
               REGION "FLASHING"
                   IF #retLogical.acutal.btn[#pBtn] THEN

                       REGION "FLASH COLOR 1"
                           IF NOT #btnParams.btn[#pBtn].flash THEN
                               IF #old.btnParam.btn[#pBtn].flash THEN
                                   #color := #btnParams.btn[#pBtn].cOn1;
                                   #draw := TRUE;
                               END_IF;
                           END_IF;
                       END_REGION

                       REGION "FLASH COLOR 2"
                           IF #btnParams.btn[#pBtn].flash THEN
                               IF NOT #old.btnParam.btn[#pBtn].flash THEN
                                   #color := #btnParams.btn[#pBtn].cOn2;
                                   #draw := TRUE;
                               END_IF;
                           END_IF;
                       END_REGION

                   END_IF;
               END_REGION

               REGION "DRAW TO BUTTON"
                   IF #draw THEN
                       #draw := FALSE;
                       "KP8 Driver: Color"(btnColor := #colorMask,
                                           btnNum := #pBtn,
                                           lblColor := #color);
                   END_IF;
               END_REGION

           END_FOR;
       END_REGION

   END_REGION

   REGION "CHANGE DETECTION"
       #old.btnParam := #btnParams;
       #old.kp8DI := #kp8DI;
       #old.logical := #retLogical.acutal;
       #old.physical := #btnPress;
   END_REGION

   REGION "OUTPUT"
       #kp8DQ := #colorMask;
       #physical := #retPhysical;
       #logical := #retLogical;
   END_REGION
END_FUNCTION_BLOCK

FUNCTION "KP8 Driver: HMI Emulator: Animation" : USInt   // FC26, SCL
{ S7_Optimized_Access := 'TRUE' }
VERSION : 0.1
   VAR_INPUT
      kp8Color : DWord;
      btnNumber : Int;
   END_VAR
   VAR_TEMP
      animate : USInt;
      blue : USInt;
      colorDWord : DWord;
      colorInt : DInt;
      green : USInt;
      off : USInt;
      red : USInt;
      white : USInt;
      yellow : USInt;
   END_VAR
   VAR CONSTANT
      blueMask : DInt := 16#0000_0100;
      btnMask : DInt := 16#0101_0100;
      greenMask : DInt := 16#0001_0000;
      offMask : DInt := 16#0000_0000;
      redMask : DInt := 16#0100_0000;
      whiteMask : DInt := 16#0101_0100;
      yellowMask : DInt := 16#0101_0000;
   END_VAR
BEGIN
   REGION "COPY TO LOCAL"
       #blue := "BLUE_LIGHT_BACKGROUND";
       #green := "GREEN_LIGHT_BACKGROUND";
       #off := "invisible";
       #red := "RED_LIGHT_BACKGROUND";
       #white := "WHITE_BACKGROUND";
       #yellow := "YELLOW_LIGHT_BACKGROUND";
   END_REGION

   REGION "ISOLATE BUTTON COLOR"
       #colorDWord := SHR_DWORD(IN := #kp8Color,N := INT_TO_ULINT(#btnNumber));
       #colorDWord := #colorDWord AND #btnMask;
       #colorInt := DWORD_TO_DINT(#colorDWord);
   END_REGION

   REGION "DETERMINE ANIMATION"
       CASE #colorInt OF
           #blueMask:
               #animate := #blue;
           #greenMask:
               #animate := #green;
           #redMask:
               #animate := #red;
           #whiteMask:
               #animate := #white;
           #yellowMask:
               #animate := #yellow;
           ELSE
               #animate := #off;
       END_CASE;
   END_REGION

   REGION "RETURN VALUE"
       #"KP8 Driver: HMI Emulator: Animation" := #animate;
   END_REGION
END_FUNCTION

FUNCTION "KP8 Driver: Group" : Void   // FC50, SCL
{ S7_Optimized_Access := 'TRUE' }
VERSION : 0.1
   VAR_INPUT
      btnNumber : Int;
      btnsParams : "KP8 Driver: Parameters: 8 Buttons";
   END_VAR
   VAR_IN_OUT
      logical : "KP8 Driver: Feedback Data";
   END_VAR
   VAR_TEMP
      pBtn : Int;
      retLogical : "KP8 Driver: Feedback Data";
      testGroup : Int;
      thisGroup : Int;
   END_VAR
BEGIN
   REGION "EXIT IF GROUP EQUALS 0"
       #thisGroup := #btnsParams.btn[#btnNumber].group;
       IF #thisGroup = 0 THEN
           RETURN;
       END_IF;
   END_REGION

   REGION "COPY TO LOCAL"
       #retLogical := #logical;
   END_REGION

   REGION "FOR EACH BUTTONS' PARAMETERS"
       FOR #pBtn := 0 TO 7 DO

           REGION "SKIP THE CURRENT BUTTON"
               IF #pBtn = #btnNumber THEN
                   GOTO NEXT;
               END_IF;
           END_REGION

           REGION "GROUP EXCLUSION"
               #testGroup := #btnsParams.btn[#pBtn].group;
               IF #testGroup = #thisGroup THEN
                   #retLogical.acutal.btn[#pBtn] := FALSE;
               END_IF;
           END_REGION

       NEXT:
           ;

       END_FOR;
   END_REGION

   REGION "OUTPUT"
       #logical := #retLogical;
   END_REGION
END_FUNCTION

FUNCTION "KP8 Driver: Toggle" : Void   // FC51, SCL
{ S7_Optimized_Access := 'TRUE' }
VERSION : 0.1
   VAR_INPUT
      signal : Bool;   // edge signal
   END_VAR
   VAR_IN_OUT
      state : Bool;   // logical button state
   END_VAR
BEGIN
   IF #signal THEN
       #state := NOT #state;
   END_IF;
END_FUNCTION

FUNCTION "KP8 Driver: Feedback" : Void   // FC52, SCL
{ S7_Optimized_Access := 'TRUE' }
VERSION : 0.1
   VAR_INPUT
      signal : Bool;
      oldSignal : Bool;
      btnNumber : Int;
   END_VAR
   VAR_IN_OUT
      feedback : "KP8 Driver: Feedback Data";
   END_VAR
   VAR_TEMP
      ret : "KP8 Driver: Feedback Data";
   END_VAR
BEGIN
   REGION "COPY TO LOCAL"
       #ret := #feedback;
       #ret.acutal.btn[#btnNumber] := #signal;
   END_REGION

   REGION "DEFAULT"
       #ret.rising.btn[#btnNumber] := FALSE;
       #ret.falling.btn[#btnNumber] := FALSE;
   END_REGION

   REGION "ON NEW INPUT"
       IF #signal <> #oldSignal THEN

           REGION "RISING EDGE"
               IF #signal AND NOT #oldSignal THEN
                   #ret.rising.btn[#btnNumber] := TRUE;
               END_IF;
           END_REGION

           REGION "FALLING EDGE"
               IF NOT #signal AND #oldSignal THEN
                   #ret.falling.btn[#btnNumber] := TRUE;
               END_IF;
           END_REGION

       END_IF;
   END_REGION


   REGION "OUTPUT"
       #feedback := #ret;
   END_REGION
END_FUNCTION

FUNCTION "KP8 Driver: State" : Void   // FC53, SCL
{ S7_Optimized_Access := 'TRUE' }
VERSION : 0.1
   VAR_INPUT
      press : "KP8 Driver: Feedback Data";
      btnNumber : Int;
      btnParams : "KP8 Driver: Parameters: 8 Buttons";
   END_VAR
   VAR_IN_OUT
      state : "KP8 Driver: Feedback Data";
   END_VAR
   VAR_TEMP
      pBtn : Int;
      retState : "KP8 Driver: Feedback Data";
   END_VAR
BEGIN
   REGION "RETURN ON INACTIVE BUTTON"
       IF NOT #btnParams.btn[#btnNumber].activate THEN
           RETURN;
       END_IF;
   END_REGION

   REGION "COPY TO LOCAL"
       #retState := #state;
   END_REGION

   REGION "MODE IS MOMENTARY"
       IF NOT #btnParams.btn[#btnNumber].mode THEN
           #retState.acutal.btn[#btnNumber] := #press.acutal.btn[#btnNumber];
       END_IF;
   END_REGION

   REGION "MAINTINED"
       IF #btnParams.btn[#btnNumber].mode THEN
           "KP8 Driver: Toggle"(signal := #press.rising.btn[#btnNumber],
                                state := #retState.acutal.btn[#btnNumber]);
       END_IF;
   END_REGION

   REGION "GROUP EXCLUSIVITY"
       IF #press.rising.btn[#btnNumber] THEN
           "KP8 Driver: Group"(btnNumber := #btnNumber,
                               btnsParams := #btnParams,
                               logical := #retState);
       END_IF;
   END_REGION

   REGION "OUTPUT"
       #state := #retState;
   END_REGION
END_FUNCTION

FUNCTION "KP8 Driver: Color" : Void   // FC54, SCL
{ S7_Optimized_Access := 'TRUE' }
VERSION : 0.1
   VAR_INPUT
      btnNum : Int;
      lblColor : String;   // 'red', 'green', 'blue', 'yellow', 'white', 'off'
   END_VAR
   VAR_IN_OUT
      btnColor : DWord;
   END_VAR
   VAR_TEMP
      btnMask : DWord;
      uColor : String;
      ret : DWord;
   END_VAR
   VAR CONSTANT
      btnMskRed : DWord := DWORD#16#0100_0000;
      btnMskGreen : DWord := DWORD#16#0001_0000;
      btnMskBlue : DWord := DWORD#16#0000_0100;
      btnMskYellow : DWord := DWORD#16#0101_0000;
      btnMskWhite : DWord := DWORD#16#0101_0100;
      btnMskOff : DWord := DWORD#16#FEFE_FEFF;
   END_VAR
BEGIN
   #ret := #btnColor;

   #ret := #ret AND ROL(IN := #btnMskOff,
                        N := INT_TO_UDINT(#btnNum));

   #uColor := #lblColor;
   "Upper"(#uColor);

   IF (#uColor = 'RED') THEN
       #btnMask := #btnMskRed;
   ELSIF (#uColor = 'GREEN') THEN
       #btnMask := #btnMskGreen;
   ELSIF (#uColor = 'BLUE') THEN
       #btnMask := #btnMskBlue;
   ELSIF (#uColor = 'YELLOW') THEN
       #btnMask := #btnMskYellow;
   ELSIF (#uColor = 'WHITE') THEN
       #btnMask := #btnMskWhite;
   ELSIF (#uColor = 'OFF') THEN
       ;
   END_IF;

   #ret := #ret OR SHL(IN := #btnMask,
                       N := INT_TO_UDINT(#btnNum));

   #btnColor := #ret;
END_FUNCTION

FUNCTION "KP8 Driver: HMI Emulator: Button Presses" : Word   // FC82, SCL
{ S7_Optimized_Access := 'TRUE' }
VERSION : 0.1
   VAR_INPUT
      pbs : DWord;
   END_VAR
   VAR_TEMP
      ret : Word;
   END_VAR
BEGIN
   #"KP8 Driver: HMI Emulator: Button Presses".%B1 := #pbs.%B0;
   #"KP8 Driver: HMI Emulator: Button Presses".%B0 := #pbs.%B1;
END_FUNCTION

// folder: Utilities

FUNCTION_BLOCK "Pulses: Button Collection"   // FB22, SCL
{ S7_Optimized_Access := 'TRUE' }
VERSION : 0.1
   VAR_INPUT
      btns : Variant;
   END_VAR
   VAR_IN_OUT
      pulses : Variant;
   END_VAR
   VAR
      old : Array[0..#u_bound] of Int;
   END_VAR
   VAR_TEMP
      eval : Array[0..#u_bound] of Int;
      i : Int;
      len_btns : UDInt;
      ret : Array[0..#u_bound] of Int;
      RET_VAL : Int;
   END_VAR
   VAR CONSTANT
      u_bound : Int := 999;
   END_VAR
BEGIN
   REGION "GET ARRAY LENGTH"
       #len_btns := CountOfElements(#btns);
   END_REGION


   REGION "COPY TO LOCAL"
       #RET_VAL := MOVE_BLK_VARIANT(SRC := #btns,
                                    COUNT := #len_btns,
                                    SRC_INDEX := 0,
                                    DEST_INDEX := 0,
                                    DEST => #eval);
   END_REGION


   REGION "CHECK FOR FALLING EDGE"
       FOR #i := 0 TO #u_bound DO
           IF #eval[#i] = 0 AND #old[#i] = 1 THEN
               #ret[#i] := 1;
           END_IF;
       END_FOR;
   END_REGION


   REGION "SAVE LAST SCAN"
       #old := #eval;
   END_REGION


   REGION "RETURN"
       #RET_VAL := MOVE_BLK_VARIANT(SRC := #ret,
                                    COUNT := #len_btns,
                                    SRC_INDEX := 0,
                                    DEST_INDEX := 0,
                                    DEST => #pulses);
   END_REGION
END_FUNCTION_BLOCK

FUNCTION_BLOCK "Push Button"   // FB41, SCL
{ S7_Optimized_Access := 'TRUE' }
VERSION : 0.1
   VAR_IN_OUT
      interface : "PB Data";
      feedback : "PB Data: State Changes";
   END_VAR
   VAR
      old : "PB Data";
   END_VAR
   VAR_TEMP
      ret : Bool;
   END_VAR
BEGIN
   REGION "ACTUATE"
       #feedback.actuate.actual := #interface.actuate;
       #feedback.actuate.rising := "Bool: Rising Edge"(signal := #interface.actuate, old_signal := #old.actuate);
       #feedback.actuate.falling := "Bool: Falling Edge"(signal := #interface.actuate, old_signal := #old.actuate);
   END_REGION

   REGION "ANIMATE"
       #feedback.animate.rising := "USInt: Value Change"(value := #interface.animate, old_value := #old.animate);
   END_REGION

   REGION "ENABLE"
       #feedback.enable.rising := "Bool: Rising Edge"(signal := #interface.enable, old_signal := #old.enable);
       #feedback.enable.actual := #interface.enable;
       #feedback.enable.falling := "Bool: Falling Edge"(signal := #interface.enable, old_signal := #old.enable);
   END_REGION

   REGION "LABEL"
       #feedback.label.rising := "WString: Value Change"(value := #interface.label, old_value := #old.label);
   END_REGION

   REGION "LIST SELECT"
       #feedback.listSelect.rising := "UInt: Value Change"(value := #interface.listSelect, old_value := #old.listSelect);
   END_REGION

   REGION "VISIBLE"
       #feedback.visible.rising := "Bool: Rising Edge"(signal := #interface.visible, old_signal := #old.visible);
       #feedback.visible.actual := #interface.visible;
       #feedback.visible.falling := "Bool: Falling Edge"(signal := #interface.visible, old_signal := #old.visible);
   END_REGION

   REGION "SAVE OLD VALUES"
       #old := #interface;
   END_REGION
END_FUNCTION_BLOCK

FUNCTION_BLOCK "IO Field"   // FB48, SCL
{ S7_Optimized_Access := 'TRUE' }
VERSION : 0.1
   VAR_IN_OUT
      interface : "IO Field Data: Label with Data";
      feedback : "IO Field: Feedback";
   END_VAR
   VAR
      old : "IO Field Data: Label with Data";
   END_VAR
BEGIN
   REGION "ANIMATE"
       #feedback.animate.rising := "USInt: Value Change"(value := #interface.animate, old_value := #old.animate);
   END_REGION

   REGION "ENABLE"
       #feedback.enable.rising := "Bool: Rising Edge"(signal := #interface.enable, old_signal := #old.enable);
       #feedback.enable.actual := #interface.enable;
       #feedback.enable.falling := "Bool: Falling Edge"(signal := #interface.enable, old_signal := #old.enable);
   END_REGION

   REGION "INPUT FINISHED"
       #feedback.input_finished.rising := "Bool: Rising Edge"(signal := #interface.input_finished, old_signal := #old.input_finished);
       #feedback.input_finished.actual := #interface.input_finished;
       #feedback.input_finished.falling := "Bool: Falling Edge"(signal := #interface.input_finished, old_signal := #old.input_finished);
   END_REGION

   REGION "VALUE CHANGED"
       #feedback.value.rising := "WString: Value Change"(value := #interface.value, old_value := #old.value);
   END_REGION

   REGION "VISIBLE"
       #feedback.visible.rising := "Bool: Rising Edge"(signal := #interface.visible, old_signal := #old.visible);
       #feedback.visible.actual := #interface.visible;
       #feedback.visible.falling := "Bool: Falling Edge"(signal := #interface.visible, old_signal := #old.visible);
   END_REGION

   REGION "SAVE OLD VALUES"
       #old := #interface;
   END_REGION
END_FUNCTION_BLOCK

FUNCTION "Animate Bool" : USInt   // FC9, SCL
{ S7_Optimized_Access := 'TRUE' }
VERSION : 0.1
   VAR_INPUT
      true_color : USInt;
      false_color : USInt;
      evaluation_signal : Bool;
   END_VAR
   VAR_TEMP
      animate : USInt;
   END_VAR
BEGIN
   REGION "FALSE COLOR"
       IF NOT #evaluation_signal THEN
           #animate := #false_color;
       END_IF;
   END_REGION

   REGION "TRUE COLOR"
       IF #evaluation_signal THEN
           #animate := #true_color;
       END_IF;
   END_REGION

   REGION "FUNCTION RETURN"
       #"Animate Bool" := #animate;
   END_REGION
END_FUNCTION

FUNCTION "Pointer Calc: KP8 Labels" : Int   // FC25, SCL
{ S7_Optimized_Access := 'TRUE' }
VERSION : 0.1
   VAR_INPUT
      index : Int;
   END_VAR
   VAR_TEMP
      val : Int;
   END_VAR
BEGIN
   IF #index >= 4 THEN
       #val := 7 - (#index - 4) * 2;
   END_IF;

   IF #index <= 3 THEN
       #val := 8 - #index * 2;
   END_IF;

   #"Pointer Calc: KP8 Labels" := #val;
END_FUNCTION

FUNCTION "Row Pointer: Roll Over" : Void   // FC33, SCL
{ S7_Optimized_Access := 'TRUE' }
VERSION : 0.1
   VAR_INPUT
      limit : Int;
   END_VAR
   VAR_IN_OUT
      pointer : Int;
   END_VAR
BEGIN
   REGION "INCREMENT"
       #pointer += 1;
   END_REGION

   REGION "HIGH LIMIT ROLLOVER"
       IF #pointer > "partReqDataRowCount" THEN
           #pointer := 0;
       END_IF;
   END_REGION
END_FUNCTION

FUNCTION "LRUD KP8 Remap" : Int   // FC35, SCL
{ S7_Optimized_Access := 'TRUE' }
VERSION : 0.1
   VAR_INPUT
      btnNum : Int;
   END_VAR
   VAR_TEMP
      output : Int;
   END_VAR
BEGIN
   IF #btnNum MOD 2 = 0 THEN
       #output := 7 - #btnNum / 2;
   END_IF;
   IF #btnNum MOD 2 <> 0 THEN
       #output := 3 - #btnNum / 2;
   END_IF;
   #"LRUD KP8 Remap" := #output;
END_FUNCTION

FUNCTION "Validate PN" : Bool   // FC42, SCL
{ S7_Optimized_Access := 'TRUE' }
VERSION : 0.1
   VAR_INPUT
      pnCode : DInt;
      pnLib : "Recipe: PN Text Library";
   END_VAR
   VAR_TEMP
      pn : WString;
      ret : Bool;
   END_VAR
BEGIN
   REGION "GET PN FROM LIBRARY"
       #pn := "Get PN From Library"(pnLib := #pnLib,
                                pnCode := #pnCode);
   END_REGION

   REGION "BUTTON HAS NO PN"
       IF LEN(#pn) = 0 THEN
           #ret := FALSE;
       END_IF;
   END_REGION

   REGION "BUTTON HAS PN"
       IF LEN(#pn) <> 0 THEN
           #ret := TRUE;
       END_IF;
   END_REGION

   REGION "RETURN"
       #"Validate PN" := #ret;
   END_REGION
END_FUNCTION

FUNCTION "Row Pointer: Post Collapse" : Void   // FC56, SCL
{ S7_Optimized_Access := 'TRUE' }
VERSION : 0.1
   VAR_INPUT
      dataTable : "Part Request Data";
   END_VAR
   VAR_IN_OUT
      pDataRow : Int;
   END_VAR
   VAR_TEMP
      pRow : Int;
   END_VAR
BEGIN
   REGION "SCAN TABLE"
       WHILE #dataTable.row[#pRow] <> -1 AND #pRow <= "partReqDataRowCount" DO
           #pRow += 1;
       END_WHILE;
   END_REGION

   REGION "TABLE NOT FULL"
       IF #pRow <="partReqDataRowCount" THEN
           #pDataRow := #pRow;
           RETURN;
       END_IF;
   END_REGION

   REGION "TABLE FULL"
       IF #pRow > "partReqDataRowCount" THEN
           #pDataRow := 0;
           RETURN;
       END_IF;
   END_REGION
END_FUNCTION

FUNCTION "Length" : UDInt   // FC60, SCL
{ S7_Optimized_Access := 'TRUE' }
VERSION : 0.1
   VAR_INPUT
      "array" : Variant;
   END_VAR
   VAR_TEMP
      status : DInt;
      ret : UDInt;
   END_VAR
BEGIN
   #ret := CountOfElements(#array);
   #Length := #ret;
END_FUNCTION

FUNCTION "Part Ordered" : Bool   // FC90, SCL
{ S7_Optimized_Access := 'TRUE' }
VERSION : 0.1
// checks state to see if the part has been ordered by the warehouse; returns a bool
   VAR_INPUT
      state : Int;
   END_VAR
   VAR_TEMP
      ret : Bool;
   END_VAR
BEGIN
   IF #state / 10 = 2 THEN
       #ret := TRUE;
   END_IF;
   #"Part Ordered" := #ret;
END_FUNCTION

FUNCTION "Is HMI Station" : Bool   // FC96, SCL
{ S7_Optimized_Access := 'TRUE' }
VERSION : 0.1
   VAR_INPUT
      stn : "Station: Single Station";
   END_VAR
   VAR_TEMP
      ret : Bool;
   END_VAR
BEGIN
   REGION "CHECK WIP COUNT"
       IF #stn.wipData.count > 0 THEN
           #ret := TRUE;
       END_IF;
   END_REGION


   REGION "RETURN"
       #"Is HMI Station" := #ret;
   END_REGION
END_FUNCTION

FUNCTION "Toggle" : Void   // FC103, SCL
{ S7_Optimized_Access := 'TRUE' }
VERSION : 0.1
   VAR_INPUT
      pulse : Bool;
   END_VAR
   VAR_IN_OUT
      state : Bool;
   END_VAR
   VAR_TEMP
      ret : Bool;
   END_VAR
BEGIN
   REGION "COPY TO LOCAL"
       #ret := #state;
   END_REGION


   REGION "TOGGLE ON PULSE"
       IF #pulse THEN
           #ret := NOT #ret;
       END_IF;
   END_REGION


   REGION "RETURN"
       #state := #ret;
   END_REGION
END_FUNCTION

FUNCTION "Count Selected Stations" : Int   // FC105, SCL
{ S7_Optimized_Access := 'TRUE' }
VERSION : 0.1
   VAR_INPUT
      selected_stns : Array[0.."STATION_COUNT"] of Bool;
   END_VAR
   VAR_TEMP
      count : Int;
      i : Int;
   END_VAR
BEGIN
   REGION "CHECK EACH STATION"
       FOR #i := 0 TO "STATION_COUNT" DO
           IF #selected_stns[#i] THEN
               #count += 1;
           END_IF;
       END_FOR;
   END_REGION


   REGION "RETURN COUNT"
       #"Count Selected Stations" := #count;
   END_REGION
END_FUNCTION

FUNCTION "Get Station Index From Id" : Int   // FC106, SCL
{ S7_Optimized_Access := 'TRUE' }
VERSION : 0.1
   VAR_INPUT
      line_name : WString;
      drop_zone : USInt;
      stns : "Station: All Stations";
   END_VAR
   VAR_TEMP
      i : Int;
      ret : Int;
   END_VAR
BEGIN
   REGION "MATCH LINE NAME AND DROP ZONE"
       FOR #i := 0 TO "STATION_COUNT" DO
           IF #line_name = #stns.stn[#i].id.lineName THEN
               IF #drop_zone = #stns.stn[#i].id.dropZone THEN
                   #ret := #i;
                   EXIT;
               END_IF;
           END_IF;
       END_FOR;
   END_REGION


   REGION "RETURN"
       #"Get Station Index From Id" := #ret;
   END_REGION
END_FUNCTION

FUNCTION "Get First Selected Station" : Int   // FC108, SCL
{ S7_Optimized_Access := 'TRUE' }
VERSION : 0.1
   VAR_INPUT
      selected_stns : Array[0.."STATION_COUNT"] of Bool;
   END_VAR
   VAR_TEMP
      eval_station_index : Int;
      i : Int;
   END_VAR
BEGIN
   REGION "FIND FIRST SELECTED STATION"
       FOR #i := 0 TO "STATION_COUNT" DO
           IF #selected_stns[#i] THEN
               #eval_station_index := #i;
               EXIT;
           END_IF;
       END_FOR;
   END_REGION


   REGION "RETURN"
       #"Get First Selected Station" := #eval_station_index;
   END_REGION
END_FUNCTION

FUNCTION "Array: Int: Fill" : Void   // FC109, SCL
{ S7_Optimized_Access := 'TRUE' }
VERSION : 0.1
   VAR_INPUT
      int_in : Int;
   END_VAR
   VAR_OUTPUT
      array_out : Variant;
   END_VAR
   VAR_TEMP
      i : Int;
      internal_array : Array[0..999] of Int;
      len_array_out : UDInt;
      status : Int;
   END_VAR
BEGIN
   REGION "GET LENGHT"
       #len_array_out := CountOfElements(#array_out);
   END_REGION


   REGION "FILL LENGTH WITH BYTE IN"
       FOR #i := 0 TO UDINT_TO_INT(#len_array_out) - 1 DO
           #internal_array[#i] := #int_in;
       END_FOR;
   END_REGION


   REGION "RETURN"
       #status := MOVE_BLK_VARIANT(SRC := #internal_array,
                                   COUNT := #len_array_out,
                                   SRC_INDEX := 0,
                                   DEST_INDEX := 0,
                                   DEST => #array_out);
   END_REGION
END_FUNCTION

FUNCTION "Array: DInt: Is Element" : Bool   // FC111, SCL
{ S7_Optimized_Access := 'TRUE' }
VERSION : 0.1
   VAR_INPUT
      array_of_int : Variant;
      search_term : DInt;
   END_VAR
   VAR_TEMP
      i : Int;
      len_as_udint : UDInt;
      len_as_int : Int;
      ret : Bool;
      status : Int;
      t_array : Array[0..#u_bound] of DInt;
   END_VAR
   VAR CONSTANT
      u_bound : Int := 999;
   END_VAR
BEGIN
   REGION "LOCAL VARIABLES"
       #len_as_udint := CountOfElements(#array_of_int);
       #len_as_int := UDINT_TO_INT(#len_as_udint) - 1;
       #status := MOVE_BLK_VARIANT(SRC := #array_of_int,
                                   COUNT := #len_as_udint,
                                   SRC_INDEX := 0,
                                   DEST_INDEX := 0,
                                   DEST => #t_array);
   END_REGION


   REGION "SEARCH ARRAY"
       FOR #i := 0 TO #len_as_int DO
           IF #t_array[#i] = #search_term THEN
               #ret := TRUE;
               EXIT;
           END_IF;
       END_FOR;
   END_REGION


   REGION "RETURN"
       #"Array: DInt: Is Element" := #ret;
   END_REGION
END_FUNCTION

FUNCTION "Get WIP Station by Global Index" : "WIP: Station"   // FC113, SCL
{ S7_Optimized_Access := 'TRUE' }
VERSION : 0.1
   VAR_INPUT
      index : Int;
      wip_stations : "Recipe: HMI Stations Saved Wips";
   END_VAR
   VAR_TEMP
      i : Int;
      ret : "WIP: Station";
   END_VAR
BEGIN
   REGION "FIND STATION"
       FOR #i := 0 TO "hmi_station_count" DO
           IF #wip_stations.stn[#i].pStn = #index THEN
               #ret := #wip_stations.stn[#i];
               EXIT;
           END_IF;
       END_FOR;
   END_REGION


   REGION "RETURN"
       #"Get WIP Station by Global Index" := #ret;
   END_REGION
END_FUNCTION

FUNCTION "Array: Int: Collapse" : Void   // FC114, SCL
{ S7_Optimized_Access := 'TRUE' }
VERSION : 0.1
   VAR_INPUT
      null_value : Int;   // value that indicates null data
   END_VAR
   VAR_IN_OUT
      int_array : Variant;
   END_VAR
   VAR_TEMP
      i : Int;
      j : Int;
      len_int : Int;
      len_udint : UDInt;
      status : Int;
      t_int_array : Array[0..999] of Int;
   END_VAR
BEGIN
   REGION "COPY TO LOCAL MEMORY"
       #len_udint := CountOfElements(#int_array);
       #len_int := UDINT_TO_INT(#len_udint) - 1;
       #status := MOVE_BLK_VARIANT(SRC := #int_array,
                                   COUNT := #len_udint,
                                   SRC_INDEX := 0,
                                   DEST_INDEX := 0,
                                   DEST => #t_int_array);
   END_REGION

   REGION "COLLAPSE IN PLACE"
       FOR #i := 0 TO #len_int - 1 DO
           IF #t_int_array[#i] = #null_value THEN
               FOR #j := #i + 1 TO #len_int DO
                   IF #t_int_array[#j] <> #null_value THEN
                       #t_int_array[#i] := #t_int_array[#j];
                       #t_int_array[#j] := #null_value;
                       EXIT;
                   END_IF;
               END_FOR;
           END_IF;
       END_FOR;
   END_REGION

   REGION "RETURN"
       #status := MOVE_BLK_VARIANT(SRC := #t_int_array,
                                   COUNT := #len_udint,
                                   SRC_INDEX := 0,
                                   DEST_INDEX := 0,
                                   DEST => #int_array);
   END_REGION
END_FUNCTION

FUNCTION "Count Collapsed Int Array" : Int   // FC115, SCL
{ S7_Optimized_Access := 'TRUE' }
VERSION : 0.1
   VAR_INPUT
      null_value : Int;
      "array" : Variant;
   END_VAR
   VAR_TEMP
      count : Int;
      i : Int;
      len_int : Int;
      len_udint : UDInt;
      status : Int;
      t_array : Array[0..999] of Int;
   END_VAR
BEGIN
   REGION "NOTES"
       (*
       returns the number of valid elements in a collapsed int array
       *)
   END_REGION


   REGION "COPY TO LOCAL"
       #len_udint := CountOfElements(#array);
       #len_int := UDINT_TO_INT(#len_udint) - 1;
       #status := MOVE_BLK_VARIANT(SRC := #array,
                                   COUNT := #len_udint,
                                   SRC_INDEX := 0,
                                   DEST_INDEX := 0,
                                   DEST => #t_array);
   END_REGION


   REGION "SCAN FOR FIRST NULL"
       FOR #i := 0 TO #len_int DO
           IF #t_array[#i] = #null_value THEN
               EXIT;
           END_IF;
           IF #t_array[#i] <> #null_value THEN
               #count += 1;
           END_IF;
       END_FOR;
   END_REGION


   REGION "RETURN"
       #"Count Collapsed Int Array" := #count;
   END_REGION
END_FUNCTION

FUNCTION "Array: Bool: List Indices of True" : Void   // FC120, SCL
{ S7_Optimized_Access := 'TRUE' }
VERSION : 0.1
   VAR_INPUT
      array_of_bool : Array[0.."STATION_COUNT"] of Bool;
   END_VAR
   VAR_OUTPUT
      list_of_indices : Variant;
   END_VAR
   VAR_TEMP
      i : Int;
      p_ret : Int;
      ret : Array[0.."STATION_COUNT"] of Int;
      status : Int;
   END_VAR
BEGIN
   REGION "FILL RETURN ARRAY"
       "Array: Int: Fill"(int_in := -1,
                        array_out => #ret);
   END_REGION


   REGION "INSERT INDICES INTO RETURN ARRAY"
       FOR #i := 0 TO "STATION_COUNT" DO
           IF #array_of_bool[#i] THEN
               #ret[#p_ret] := #i;
               #p_ret += 1;
           END_IF;
       END_FOR;
   END_REGION


   REGION "RETURN"
       #status := MOVE_BLK_VARIANT(SRC := #ret,
                                   COUNT := INT_TO_UDINT("STATION_COUNT"),
                                   SRC_INDEX := 0,
                                   DEST_INDEX := 0,
                                   DEST => #list_of_indices);
   END_REGION
END_FUNCTION

FUNCTION "Array: Int: Is Element" : Bool   // FC121, SCL
{ S7_Optimized_Access := 'TRUE' }
VERSION : 0.1
   VAR_INPUT
      array_of_int : Variant;
      search_term : Int;
   END_VAR
   VAR_TEMP
      i : Int;
      len_as_udint : UDInt;
      len_as_int : Int;
      ret : Bool;
      status : Int;
      t_array : Array[0..999] of Int;
   END_VAR
BEGIN
   REGION "LOCAL VARIABLES"
       #len_as_udint := CountOfElements(#array_of_int);
       #len_as_int := UDINT_TO_INT(#len_as_udint) - 1;
       #status := MOVE_BLK_VARIANT(SRC := #array_of_int,
                                   COUNT := #len_as_udint,
                                   SRC_INDEX := 0,
                                   DEST_INDEX := 0,
                                   DEST => #t_array);
   END_REGION


   REGION "SEARCH ARRAY"
       FOR #i := 0 TO #len_as_int DO
           IF #t_array[#i] = #search_term THEN
               #ret := TRUE;
               EXIT;
           END_IF;
       END_FOR;
   END_REGION


   REGION "RETURN"
       #"Array: Int: Is Element" := #ret;
   END_REGION
END_FUNCTION

FUNCTION "Remap Int Array" : Void   // FC122, SCL
{ S7_Optimized_Access := 'TRUE' }
VERSION : 0.1
   VAR_INPUT
      source_int_array : Variant;
   END_VAR
   VAR_IN_OUT
      destination_int_array : Variant;
   END_VAR
   VAR_TEMP
      len_destination : UDInt;
      status : Int;
   END_VAR
BEGIN
   #len_destination := CountOfElements(#destination_int_array);
   #status := MOVE_BLK_VARIANT(SRC := #source_int_array,
                               COUNT := #len_destination,
                               SRC_INDEX := 0,
                               DEST_INDEX := 0,
                               DEST => #destination_int_array);
END_FUNCTION

FUNCTION "Count Selected WIPs" : Int   // FC126, SCL
{ S7_Optimized_Access := 'TRUE' }
VERSION : 0.1
   VAR_INPUT
      selected_WIPs : Array[0.."wipCount"] of DInt;
   END_VAR
   VAR_TEMP
      count : Int;
      i : Int;
   END_VAR
BEGIN
   REGION "CHECK EACH STATION"
       FOR #i := 0 TO "wipCount" DO
           IF #selected_WIPs[#i] = INT_TO_DINT("NULL_TOKEN") THEN
               EXIT;
           END_IF;
           IF #selected_WIPs[#i] <> INT_TO_DINT("NULL_TOKEN") THEN
               #count += 1;
           END_IF;
       END_FOR;
   END_REGION


   REGION "RETURN COUNT"
       #"Count Selected WIPs" := #count;
   END_REGION
END_FUNCTION

FUNCTION "Count Selected Buttons" : Int   // FC127, SCL
{ S7_Optimized_Access := 'TRUE' }
VERSION : 0.1
   VAR_INPUT
      selected_buttons : Array[0.."STATION_BUTTON_COUNT"] of Bool;
   END_VAR
   VAR_TEMP
      count : Int;
      i : Int;
   END_VAR
BEGIN
   REGION "CHECK EACH STATION"
       FOR #i := 0 TO "STATION_BUTTON_COUNT" DO
           IF #selected_buttons[#i] THEN
               #count += 1;
           END_IF;
       END_FOR;
   END_REGION


   REGION "RETURN COUNT"
       #"Count Selected Buttons" := #count;
   END_REGION
END_FUNCTION

FUNCTION "Get WIP Station Index by Global Index" : Int   // FC130, SCL
{ S7_Optimized_Access := 'TRUE' }
VERSION : 0.1
   VAR_INPUT
      global_index : Int;
      saved_WIPs : "Recipe: HMI Stations Saved Wips";
   END_VAR
   VAR_TEMP
      i : Int;
      ret : Int;
   END_VAR
BEGIN
   REGION "SEARCH FOR INDEX"
       #ret := "NULL_TOKEN";
       FOR #i := 0 TO "hmi_station_count" DO
           IF #saved_WIPs.stn[#i].pStn = #global_index THEN
               #ret := #i;
               EXIT;
           END_IF;
       END_FOR;
   END_REGION


   REGION "RETURN"
       #"Get WIP Station Index by Global Index" := #ret;
   END_REGION
END_FUNCTION

FUNCTION "Fill DInt Array" : Void   // FC131, SCL
{ S7_Optimized_Access := 'TRUE' }
VERSION : 0.1
   VAR_INPUT
      int_in : DInt;
   END_VAR
   VAR_OUTPUT
      array_out : Variant;
   END_VAR
   VAR_TEMP
      i : Int;
      internal_array : Array[0..999] of DInt;
      len_array_out : UDInt;
      status : Int;
   END_VAR
BEGIN
   REGION "GET LENGHT"
       #len_array_out := CountOfElements(#array_out);
   END_REGION


   REGION "FILL LENGTH WITH BYTE IN"
       FOR #i := 0 TO UDINT_TO_INT(#len_array_out) - 1 DO
           #internal_array[#i] := #int_in;
       END_FOR;
   END_REGION


   REGION "RETURN"
       #status := MOVE_BLK_VARIANT(SRC := #internal_array,
                                   COUNT := #len_array_out,
                                   SRC_INDEX := 0,
                                   DEST_INDEX := 0,
                                   DEST => #array_out);
   END_REGION
END_FUNCTION

FUNCTION "Collapse DInt Array" : Void   // FC132, SCL
{ S7_Optimized_Access := 'TRUE' }
VERSION : 0.1
   VAR_INPUT
      null_value : DInt;   // value that indicates null data
   END_VAR
   VAR_IN_OUT
      int_array : Variant;
   END_VAR
   VAR_TEMP
      i : Int;
      j : Int;
      len_int : Int;
      len_udint : UDInt;
      status : Int;
      t_int_array : Array[0..999] of DInt;
   END_VAR
BEGIN
   REGION "COPY TO LOCAL MEMORY"
       #len_udint := CountOfElements(#int_array);
       #len_int := UDINT_TO_INT(#len_udint) - 1;
       #status := MOVE_BLK_VARIANT(SRC := #int_array,
                                   COUNT := #len_udint,
                                   SRC_INDEX := 0,
                                   DEST_INDEX := 0,
                                   DEST => #t_int_array);
   END_REGION

   REGION "COLLAPSE IN PLACE"
       FOR #i := 0 TO #len_int - 1 DO
           IF #t_int_array[#i] = #null_value THEN
               FOR #j := #i + 1 TO #len_int DO
                   IF #t_int_array[#j] <> #null_value THEN
                       #t_int_array[#i] := #t_int_array[#j];
                       #t_int_array[#j] := #null_value;
                       EXIT;
                   END_IF;
               END_FOR;
           END_IF;
       END_FOR;
   END_REGION

   REGION "RETURN"
       #status := MOVE_BLK_VARIANT(SRC := #t_int_array,
                                   COUNT := #len_udint,
                                   SRC_INDEX := 0,
                                   DEST_INDEX := 0,
                                   DEST => #int_array);
   END_REGION
END_FUNCTION

FUNCTION "Count Collapsed DInt Array" : Int   // FC133, SCL
{ S7_Optimized_Access := 'TRUE' }
VERSION : 0.1
   VAR_INPUT
      null_value : DInt;
      "array" : Variant;
   END_VAR
   VAR_TEMP
      count : Int;
      i : Int;
      len_int : Int;
      len_udint : UDInt;
      status : Int;
      t_array : Array[0..999] of DInt;
   END_VAR
BEGIN
   REGION "NOTES"
       (*
       returns the number of valid elements in a collapsed int array
       *)
   END_REGION


   REGION "COPY TO LOCAL"
       #len_udint := CountOfElements(#array);
       #len_int := UDINT_TO_INT(#len_udint) - 1;
       #status := MOVE_BLK_VARIANT(SRC := #array,
                                   COUNT := #len_udint,
                                   SRC_INDEX := 0,
                                   DEST_INDEX := 0,
                                   DEST => #t_array);
   END_REGION


   REGION "SCAN FOR FIRST NULL"
       FOR #i := 0 TO #len_int DO
           IF #t_array[#i] = INT_TO_DINT("NULL_TOKEN") THEN
               EXIT;
           END_IF;
           IF #t_array[#i] <> #null_value THEN
               #count += 1;
           END_IF;
       END_FOR;
   END_REGION


   REGION "RETURN"
       #"Count Collapsed DInt Array" := #count;
   END_REGION
END_FUNCTION

FUNCTION "Map WIP Codes to DInt Array" : Void   // FC139, SCL
{ S7_Optimized_Access := 'TRUE' }
VERSION : 0.1
   VAR_INPUT
      station : "WIP: Station";
   END_VAR
   VAR_IN_OUT
      WIP_array : Array[0.."wipCount"] of DInt;
   END_VAR
   VAR_TEMP
      i : Int;
   END_VAR
BEGIN
   FOR #i := 0 TO "wipCount" DO
       IF #station.wip[#i].wip.code = "NULL_TOKEN" THEN
           EXIT;
       END_IF;
       #WIP_array[#i] := #station.wip[#i].wip.code;
   END_FOR;
END_FUNCTION

FUNCTION "Array: Int: Search" : Int   // FC140, SCL
{ S7_Optimized_Access := 'TRUE' }
VERSION : 0.1
   VAR_INPUT
      array_of_int : Variant;   // max upper bound 999
      search_term : Int;
   END_VAR
   VAR_TEMP
      i : Int;
      len_as_udint : UDInt;
      len_as_int : Int;
      ret : Int;
      status : Int;
      t_array : Array[0..999] of Int;
   END_VAR
   // Ret_Val : index of search term. returns -1 if not found.
BEGIN
   REGION "LOCAL VARIABLES"
       #len_as_udint := CountOfElements(#array_of_int);
       #len_as_int := UDINT_TO_INT(#len_as_udint) - 1;
       #status := MOVE_BLK_VARIANT(SRC := #array_of_int,
                                   COUNT := #len_as_udint,
                                   SRC_INDEX := 0,
                                   DEST_INDEX := 0,
                                   DEST => #t_array);
       #ret := -1;
   END_REGION


   REGION "SEARCH ARRAY"
       FOR #i := 0 TO #len_as_int DO
           IF #t_array[#i] = #search_term THEN
               #ret := #i;
               EXIT;
           END_IF;
       END_FOR;
   END_REGION


   REGION "RETURN"
       #"Array: Int: Search" := #ret;
   END_REGION
END_FUNCTION

FUNCTION "Array: Int: Intersect" : Void   // FC141, SCL
{ S7_Optimized_Access := 'TRUE' }
VERSION : 0.1
   VAR_INPUT
      "a" : Variant;   // should be array of int, max 999
      "b" : Variant;   // should be array of int, max 999
      null_value : Int;
   END_VAR
   VAR_OUTPUT
      intersect_array : Variant;   // should be array of int, max 999
   END_VAR
   VAR_TEMP
      i : Int;
      j : Int;
      len_a : Struct
         as_udint : UDInt;
         as_int : Int;
      END_STRUCT;
      len_b : Struct
         as_udint : UDInt;
         as_int : Int;
      END_STRUCT;
      len_longer : Struct
         as_udint : UDInt;
         as_int : Int;
      END_STRUCT;
      len_shorter : Struct
         as_udint : UDInt;
         as_int : Int;
      END_STRUCT;
      t_a : Array[0..#u_bound] of Int;
      p_ret : Int;
      ret : Array[0..#u_bound_double] of Int;
      t_b : Array[0..#u_bound] of Int;
      status : Int;
   END_VAR
   VAR CONSTANT
      u_bound : Int := 999;
      u_bound_double : Int := 1999;
   END_VAR
BEGIN
   REGION "GET LENGTHS"
       #len_a.as_udint := CountOfElements(#a);
       #len_a.as_int := UDINT_TO_INT(#len_a.as_udint) - 1;
       #len_b.as_udint := CountOfElements(#b);
       #len_b.as_int := UDINT_TO_INT(#len_b.as_udint) - 1;
   END_REGION

   REGION "MOVE"
       #status := MOVE_BLK_VARIANT(SRC := #a, COUNT := #len_a.as_udint, SRC_INDEX := 0, DEST_INDEX := 0, DEST => #t_a);
       #status := MOVE_BLK_VARIANT(SRC := #b, COUNT := #len_b.as_udint, SRC_INDEX := 0, DEST_INDEX := 0, DEST => #t_b);
   END_REGION

   REGION "FIND INTERSECT"
       FOR #i := 0 TO #len_a.as_int DO
           IF #t_a[#i] = #null_value THEN
               EXIT;
           END_IF;
           FOR #j := 0 TO #len_b.as_int DO
               IF #t_b[#j] = #null_value THEN
                   EXIT;
               END_IF;
               IF #t_a[#i] = #t_b[#j] THEN
                   #ret[#p_ret] := #t_a[#i];
                   #p_ret += 1;
                   EXIT;
               END_IF;
           END_FOR;
       END_FOR;
   END_REGION

   REGION "RETURN"
       #status := MOVE_BLK_VARIANT(SRC := #ret, COUNT := INT_TO_UDINT(#p_ret - 1), SRC_INDEX := 0, DEST_INDEX := 0, DEST => #intersect_array);
   END_REGION
END_FUNCTION

FUNCTION "Map Selected Stations to Int Array" : Void   // FC142, SCL
{ S7_Optimized_Access := 'TRUE' }
VERSION : 0.1
   VAR_INPUT
      selected_stations : "Selected Stations";
   END_VAR
   VAR_OUTPUT
      selected_stations_indicies : Array[0.."STATION_COUNT"] of Int;
   END_VAR
   VAR_TEMP
      i : Int;
      p_ret : Int;
      ret : Array[0.."STATION_COUNT"] of Int;
   END_VAR
BEGIN
   "Array: Int: Fill"(int_in := "NULL_TOKEN",
                      array_out => #ret);
   FOR #i := 0 TO "STATION_COUNT" DO
       IF #selected_stations.stns[#i] THEN
           #ret[#p_ret] := #i;
           #p_ret += 1;
       END_IF;
   END_FOR;
   #selected_stations_indicies := #ret;
END_FUNCTION

FUNCTION "Array: DInt: Get Index of First Occurance" : Int   // FC143, SCL
{ S7_Optimized_Access := 'TRUE' }
VERSION : 0.1
   VAR_INPUT
      dint_array : Variant;
      search_term : DInt;
   END_VAR
   VAR_TEMP
      i : Int;
      len : UDInt;
      status : Int;
      t_dint_array : Array[0..#u_bound] of DInt;
   END_VAR
   VAR CONSTANT
      u_bound : Int := 999;
   END_VAR
BEGIN
   REGION "NOTES"
       (* 
       This function returns the first occurance of the null value given 
       at the input "null_value".
       This function is commonly used on collapsed arrays.
       See "Array: DInt: Collapse" for collapse functionality.
       *)
   END_REGION


   REGION "GET LENGTH OF INPUT ARRAY"
       #len := CountOfElements(#dint_array);
       #status := MOVE_BLK_VARIANT(SRC := #dint_array, COUNT := #len, SRC_INDEX := 0, DEST_INDEX := 0, DEST => #t_dint_array);
   END_REGION


   REGION "FIND FIRST NULL, -1 IF NONE"
       (*
       Its worth noting that "Array: Dint: Is Element" could return the index of the search term
       as an output, saving the processor some work. 
       The design decision was made to re-do this work so that the functions could return their values
       insead of making use of outputs or in/outs.
       This allows for easier "in-line" use and less cluttered interfaces.
       Additionally the time complexity for "Array: DInt" Get Index of First Occurance" remains O(n).
       *)
       IF "Array: DInt: Is Element"(array_of_int := #t_dint_array, search_term := #search_term) THEN
           // the length check is left as a redundancy
           WHILE #t_dint_array[#i] <> #search_term AND INT_TO_UDINT(#i) < #len DO
               #i += 1;
           END_WHILE;
       END_IF;
   END_REGION


   REGION _name_
       #"Array: DInt: Get Index of First Occurance" := #i;
   END_REGION
END_FUNCTION

FUNCTION "Array: DInt: Intersect Exists" : Bool   // FC144, SCL
{ S7_Optimized_Access := 'TRUE' }
VERSION : 0.1
   VAR_INPUT
      "a" : Variant;   // should be array of dint, max 999
      "b" : Variant;   // should be array of dint, max 999
      null_value : DInt;
   END_VAR
   VAR_TEMP
      i : Int;
      j : Int;
      len_a : Struct
         as_udint : UDInt;
         as_int : Int;
      END_STRUCT;
      len_b : Struct
         as_udint : UDInt;
         as_int : Int;
      END_STRUCT;
      t_a : Array[0..#u_bound] of DInt;
      p_ret : Int;
      ret : Bool;
      t_b : Array[0..#u_bound] of DInt;
      status : Int;
   END_VAR
   VAR CONSTANT
      u_bound : Int := 999;
   END_VAR
BEGIN
   REGION "GET LENGHTS"
       #len_a.as_udint := CountOfElements(#a);
       #len_a.as_int := UDINT_TO_INT(#len_a.as_udint) - 1;
       #len_b.as_udint := CountOfElements(#b);
       #len_b.as_int := UDINT_TO_INT(#len_b.as_udint) - 1;
   END_REGION

   REGION "PERFORM MOVES"
       #status := MOVE_BLK_VARIANT(SRC := #a, COUNT := #len_a.as_udint, SRC_INDEX := 0, DEST_INDEX := 0, DEST => #t_a);
       #status := MOVE_BLK_VARIANT(SRC := #b, COUNT := #len_b.as_udint, SRC_INDEX := 0, DEST_INDEX := 0, DEST => #t_b);
   END_REGION


   REGION "SEARCH FOR ANY MATCHING ELEMENT"
       FOR #i := 0 TO #len_a.as_int DO

           REGION "SKIP NULL VALUES"
               IF #t_a[#i] = #null_value THEN
                   CONTINUE;
               END_IF;
           END_REGION

           REGION "INNER LOOP"
               FOR #j := 0 TO #len_b.as_int DO

                   REGION "SKIP NULL VALUES"
                       IF #t_b[#j] = #null_value THEN
                           CONTINUE;
                       END_IF;
                   END_REGION

                   REGION "SET RETURN VALUE ON MATCH"
                       IF #t_a[#i] = #t_b[#j] THEN
                           #ret := TRUE;
                           EXIT;
                       END_IF;
                   END_REGION

               END_FOR;
           END_REGION

           REGION "EXIT OUTTER LOOP IF MATCH FOUND"
               IF #ret THEN
                   EXIT;
               END_IF;
           END_REGION

       END_FOR;
   END_REGION

   REGION "RETURN"
       #"Array: DInt: Intersect Exists" := #ret;
   END_REGION
END_FUNCTION

FUNCTION "Array: DInt: Intersect" : Void   // FC145, SCL
{ S7_Optimized_Access := 'TRUE' }
VERSION : 0.1
   VAR_INPUT
      "a" : Variant;   // should be array of dint, max 999
      "b" : Variant;   // should be array of dint, max 999
      null_value : DInt;
   END_VAR
   VAR_OUTPUT
      intersect_array : Variant;   // should be array of dint, max 999
   END_VAR
   VAR_TEMP
      i : Int;
      j : Int;
      len_a : Struct
         as_udint : UDInt;
         as_int : Int;
      END_STRUCT;
      len_b : Struct
         as_udint : UDInt;
         as_int : Int;
      END_STRUCT;
      t_a : Array[0..#u_bound] of DInt;
      p_ret : Int;
      ret : Array[0..#u_bound_double] of DInt;
      t_b : Array[0..#u_bound] of DInt;
      status : Int;
   END_VAR
   VAR CONSTANT
      u_bound : Int := 999;
      u_bound_double : Int := 1999;
   END_VAR
BEGIN
   REGION "GET LENGTHS"
       #len_a.as_udint := CountOfElements(#a);
       #len_a.as_int := UDINT_TO_INT(#len_a.as_udint) - 1;
       #len_b.as_udint := CountOfElements(#b);
       #len_b.as_int := UDINT_TO_INT(#len_b.as_udint) - 1;
   END_REGION

   REGION "MOVE"
       #status := MOVE_BLK_VARIANT(SRC := #a, COUNT := #len_a.as_udint, SRC_INDEX := 0, DEST_INDEX := 0, DEST => #t_a);
       #status := MOVE_BLK_VARIANT(SRC := #b, COUNT := #len_b.as_udint, SRC_INDEX := 0, DEST_INDEX := 0, DEST => #t_b);
   END_REGION

   REGION "FIND INTERSECT"
       FOR #i := 0 TO #len_a.as_int DO
           IF #t_a[#i] = #null_value THEN
               EXIT;
           END_IF;
           FOR #j := 0 TO #len_b.as_int DO
               IF #t_b[#j] = #null_value THEN
                   EXIT;
               END_IF;
               IF #t_a[#i] = #t_b[#j] THEN
                   #ret[#p_ret] := #t_a[#i];
                   #p_ret += 1;
                   EXIT;
               END_IF;
           END_FOR;
       END_FOR;
   END_REGION

   REGION "RETURN"
       #status := MOVE_BLK_VARIANT(SRC := #ret, COUNT := INT_TO_UDINT(#p_ret - 1), SRC_INDEX := 0, DEST_INDEX := 0, DEST => #intersect_array);
   END_REGION
END_FUNCTION

FUNCTION "Bool: Rising Edge" : Bool   // FC177, SCL
{ S7_Optimized_Access := 'TRUE' }
VERSION : 0.1
   VAR_INPUT
      signal : Bool;
      old_signal : Bool;
   END_VAR
BEGIN
   #"Bool: Rising Edge" := #signal AND NOT #old_signal;
END_FUNCTION

FUNCTION "Bool: Falling Edge" : Bool   // FC178, SCL
{ S7_Optimized_Access := 'TRUE' }
VERSION : 0.1
   VAR_INPUT
      signal : Bool;
      old_signal : Bool;
   END_VAR
BEGIN
   #"Bool: Falling Edge" := NOT #signal AND #old_signal;
END_FUNCTION

FUNCTION "Int: Value Change" : Bool   // FC179, SCL
{ S7_Optimized_Access := 'TRUE' }
VERSION : 0.1
   VAR_INPUT
      value : Int;
      old_value : Int;
   END_VAR
BEGIN
   #"Int: Value Change" := #value <> #old_value;
END_FUNCTION

FUNCTION "USInt: Value Change" : Bool   // FC181, SCL
{ S7_Optimized_Access := 'TRUE' }
VERSION : 0.1
   VAR_INPUT
      value : USInt;
      old_value : USInt;
   END_VAR
BEGIN
   #"USInt: Value Change" := #value <> #old_value;
END_FUNCTION

FUNCTION "WString: Value Change" : Bool   // FC182, SCL
{ S7_Optimized_Access := 'TRUE' }
VERSION : 0.1
   VAR_INPUT
      value : WString;
      old_value : WString;
   END_VAR
BEGIN
   #"WString: Value Change" := #value <> #old_value;
END_FUNCTION

FUNCTION "UInt: Value Change" : Bool   // FC183, SCL
{ S7_Optimized_Access := 'TRUE' }
VERSION : 0.1
   VAR_INPUT
      value : UInt;
      old_value : UInt;
   END_VAR
BEGIN
   #"UInt: Value Change" := #value <> #old_value;
END_FUNCTION

// folder: Utilities/Address

FUNCTION "Address: Get Button" : DInt   // FC21, SCL
{ S7_Optimized_Access := 'TRUE' }
VERSION : 0.1
   VAR_INPUT
      address : DInt;
   END_VAR
BEGIN
   #"Address: Get Button" := #address MOD 10;
END_FUNCTION

FUNCTION "Address: Get Station" : DInt   // FC24, SCL
{ S7_Optimized_Access := 'TRUE' }
VERSION : 0.1
   VAR_INPUT
      address : DInt;
   END_VAR
BEGIN
   #"Address: Get Station" := #address / 10_000;
END_FUNCTION

FUNCTION "Address: Set Address" : DInt   // FC32, SCL
{ S7_Optimized_Access := 'TRUE' }
VERSION : 0.1
   VAR_INPUT
      pBtn : Int;
      pStn : Int;
      pWip : Int;
   END_VAR
BEGIN
   #"Address: Set Address" := INT_TO_DINT(#pStn) * 10_000 + INT_TO_DINT(#pWip) * 10 + INT_TO_DINT(#pBtn);
END_FUNCTION

FUNCTION "Address: Get Wip" : DInt   // FC88, SCL
{ S7_Optimized_Access := 'TRUE' }
VERSION : 0.1
   VAR_INPUT
      address : DInt;
   END_VAR
BEGIN
   #"Address: Get Wip" := #address - "Address: Get Station"(#address) * 10_000 - "Address: Get Button"(#address);
END_FUNCTION

// folder: Utilities/Encoding

FUNCTION "Part Number: Parse Code" : Void   // FC34, SCL
{ S7_Optimized_Access := 'TRUE' }
VERSION : 0.1
   VAR_INPUT
      code : DInt;
   END_VAR
   VAR_OUTPUT
      code_left : DInt;
      code_right : DInt;
   END_VAR
BEGIN
   IF #code > 0 THEN
       #code_left := #code / 1000;
       #code_right := #code - #code / 1000 * 1000;
   ELSE
       #code_left := 0;
       #code_right := 0;
   END_IF;
END_FUNCTION

FUNCTION "Get PN From Library" : WString   // FC37, SCL
{ S7_Optimized_Access := 'TRUE' }
VERSION : 0.1
   VAR_INPUT
      pnLib : "Recipe: PN Text Library";
      pnCode : DInt;
   END_VAR
   VAR_TEMP
      pnLeft : DInt;
      pnRight : DInt;
      output : WString;
   END_VAR
   VAR CONSTANT
      newLine : WString := WSTRING#'$L';
   END_VAR
BEGIN
   REGION "PARSE CODE"
       "Part Number: Parse Code"(code := #pnCode,
                                 code_left => #pnLeft,
                                 code_right => #pnRight);
   END_REGION

   REGION "SINGLE LINE PN"
       IF "Part Number: Is Single"(#pnCode) THEN
           #output := #pnLib.pnText[#pnLeft];
       END_IF;
   END_REGION

   REGION "DOUBLE LINE PN"
       IF "Part Number: Is Double"(#pnCode) THEN
           #output := CONCAT_WSTRING(IN1 := #pnLib.pnText[#pnLeft],
                                     IN2 := #newLine,
                                     IN3 := #pnLib.pnText[#pnRight]);
       END_IF;
   END_REGION

   REGION "OUTPUT"
       #"Get PN From Library" := #output;
   END_REGION
END_FUNCTION

